(* Logix 5000 project; controller MV vendor 1 type 14 code 217 rev 31.11; software revision 31.00; part 52 of 53 *)
(* tags used below, declared in another part *)
   Alarm_Reset : BOOL;
   CWD : CHECKWORD_FLAGS;
   Default_Check_Time : DINT;
   Dummy : BOOL;
   Item_Faults_Are_Latched : BOOL;
   Item_Simulation_Flag : BOOL;
   Mike_050419 : BOOL;
   MV_data_file_address : INT;
   MV_data_file_value_to_move : DINT;
   MV_MV20R : PlantItem;   // MV20R
   MV_MV20R_ALARM : ALARM_DIGITAL;
   MV_MV20R_D : ALIAS FOR Remote_IO:14:O.Data.9;   // Rouser drive MV20
   MV_MV20R_R : ALIAS FOR Remote_IO:15:I.Data.25;   // MV20 Rouser running signal
   MV_MV21R : PlantItem;   // MV21R
   MV_MV21R_ALARM : ALARM_DIGITAL;
   MV_MV21R_D : ALIAS FOR Remote_IO:14:O.Data.10;   // Rouser drive MV21
   MV_MV21R_R : ALIAS FOR Remote_IO:15:I.Data.26;   // MV21 Rouser running signal
   MV_MV22R : PlantItem;   // MV22R
   MV_MV22R_ALARM : ALARM_DIGITAL;
   MV_MV22R_D : ALIAS FOR Remote_IO:14:O.Data.11;   // Rouser drive MV22
   MV_MV22R_R : ALIAS FOR Remote_IO:15:I.Data.27;   // MV22 Rouser running signal
   MV_MV23R : PlantItem;   // MV23R
   MV_MV23R_ALARM : ALARM_DIGITAL;
   MV_MV23R_D : ALIAS FOR Remote_IO:14:O.Data.12;   // Rouser drive MV23
   MV_MV23R_R : ALIAS FOR Remote_IO:15:I.Data.28;   // MV23 Rouser running signal
   MV_MV35R : PlantItem;   // MV35R
   MV_MV35R_ALARM : ALARM_DIGITAL;
   MV_MV35R_D : ALIAS FOR Remote_IO:14:O.Data.8;   // Rouser drive MV35
   MV_MV35R_R : ALIAS FOR Remote_IO:15:I.Data.24;   // MV35 Rouser running signal
   MV_N101 : INT[255];   // AT INT Fermentation control integer workspace
   MV_N105 : INT[255];   // ROUSE_CTRL Rouser control progr am working regs
   MV_N105_0_1_Output_Bit : BOOL;
   MV_N105_0_6_Output_Bit : BOOL;
   MV_N105_0_7_Output_Bit : BOOL;
   MV_N105_0_8_Output_Bit : BOOL;
   MV_N106 : INT[255];   // ROUSE_BUFF Rouser control vesse l data buffer
   MV_N110 : INT[255];   // MV DATA 0 CURRENT FV DATA
   MV_N111 : INT[50];   // MV 1, CURRENT FV DATA
   MV_N112 : INT[50];   // MV 2, CURRENT FV DATA
   MV_N113 : INT[50];   // MV 3, CURRENT FV DATA
   MV_N114 : INT[50];   // MV 4, CURRENT FV DATA
   MV_N115 : INT[50];   // MV 5, CURRENT FV DATA
   MV_N116 : INT[50];   // MV 6, CURRENT FV DATA
   MV_N117 : INT[50];   // MV 7, CURRENT FV DATA
   MV_N118 : INT[50];   // MV 8, CURRENT FV DATA
   MV_N119 : INT[50];   // MV 9, CURRENT FV DATA
   MV_N12 : INT[255];   // SYS_PARMS System Parameter Fil e
   MV_N120 : INT[50];   // MV 10, CURRENT FV DATA
   MV_N121 : INT[50];   // MV 11, CURRENT FV DATA
   MV_N122 : INT[50];   // MV 12, CURRENT FV DATA
   MV_N123 : INT[50];   // MV 13, CURRENT FV DATA
   MV_N124 : INT[50];   // MV 14, CURRENT FV DATA
   MV_N125 : INT[50];   // MV 15, CURRENT FV DATA
   MV_N126 : INT[50];   // MV 16, CURRENT FV DATA
   MV_N127 : INT[50];   // MV 17, CURRENT FV DATA
   MV_N128 : INT[50];   // MV 18, CURRENT FV DATA
   MV_N129 : INT[50];   // MV 19, CURRENT FV DATA
   MV_N130 : INT[50];   // MV 30, CURRENT FV DATA
   MV_N131 : INT[50];   // MV 31, CURRENT FV DATA
   MV_N132 : INT[50];   // MV 32, CURRENT FV DATA
   MV_N133 : INT[50];   // MV 33, CURRENT FV DATA
   MV_N134 : INT[50];   // MV 34, CURRENT FV DATA
   MV_N135 : INT[50];   // MV 35, CURRENT FV DATA
   MV_N136 : INT[50];   // MV 20, CURRENT FV DATA
   MV_N137 : INT[50];   // MV 21, CURRENT FV DATA
   MV_N138 : INT[50];   // MV 22, CURRENT FV DATA
   MV_N139 : INT[50];   // MV 23, CURRENT FV DATA
   MV_N140 : INT[50];   // MV 36, CURRENT FV DATA
   MV_N141 : INT[50];   // MV 37, CURRENT FV DATA
   MV_N142 : INT[50];   // MV 38, CURRENT FV DATA
   MV_N143 : INT[50];   // MV 39, CURRENT FV DATA
   MV_N144 : INT[50];   // MV 40, CURRENT FV DATA
   MV_N145 : INT[50];   // MV 41, CURRENT FV DATA
   MV_N146 : INT[50];   // MV 42, CURRENT FV DATA
   MV_N147 : INT[50];   // MV 43, CURRENT FV DATA
   MV_N148 : INT[50];   // MV 44, CURRENT FV DATA
   MV_N149 : INT[50];   // MV 45, CURRENT FV DATA
   MV_N150 : INT[50];   // MV 36, CURRENT FV DATA
   MV_N151 : INT[50];   // MV 47, CURRENT FV DATA
   MV_SFile : INT[255];   // SLC Equivalent System File, So Original Code Can Remain
   MV_T4 : TIMER[20];
   MV_value_to_set : INT;
   MV_word_offset : INT;
   One_Second_One_Scan : ALIAS FOR One_Second_1_scan;
   Scada_Pump_Fault_No : DINT;
   Scada_Pump_H_Fault_No : DINT;
   Scada_Pump_T_Fault_No : DINT;
   Unused_Healthy_Feedback : BOOL;
   Unused_NotTripped_Feedback : BOOL;
(* MV_Common, continued *)

   24: [NEQ(MV_MV35R.DriveBits,0) OTE(MV_MV35R.CW.[CWD.AUTODRV]) ,[XIC(MV_MV35R.CW.[CWD.AUTODRV]) XIO(MV_MV35R.CW.[CWD.MANUAL]) ,XIC(MV_MV35R.CW.[CWD.MANDRV]) XIC(MV_MV35R.CW.[CWD.MANUAL]) ] OTE(MV_MV35R.CW.[CWD.OUTPUT]) ,XIC(MV_MV35R.CW.[CWD.OUTPUT]) OTE(MV_MV35R_D) ,XIC(S:FS) [OTU(MV_MV35R.CW.[CWD.MANUAL]) ,LEQ(MV_MV35R.CheckTime,0) MOV(Default_Check_Time,MV_MV35R.CheckTime) ] ,[[XIC(MV_MV35R_R) XIO(Item_Simulation_Flag) ,XIC(Item_Simulation_Flag) [XIC(MV_MV35R.CW.[CWD.OUTPUT]) XIO(MV_MV35R.CW.[CWD.SIMFAIL]) ,XIO(MV_MV35R.CW.[CWD.OUTPUT]) XIC(MV_MV35R.CW.[CWD.SIMFAIL]) ] ] OTE(MV_MV35R.CW.[CWD.RUNFB]) ,[XIC(Item_Simulation_Flag) ,XIC(MV_MV35R.CW.[CWD.CHECKOFF]) ,XIC(Unused_Healthy_Feedback) ] OTE(MV_MV35R.CW.[CWD.HEALTHYFB]) ,[XIC(Item_Simulation_Flag) ,XIC(MV_MV35R.CW.[CWD.CHECKOFF]) ,XIC(Unused_NotTripped_Feedback) ] OTE(MV_MV35R.CW.[CWD.NOTTRIPPEDFB]) ] ,[XIC(MV_MV35R.CW.[CWD.AUTODRV]) XIO(MV_MV35R.CW.[CWD.PREVSCAN]) ,XIO(MV_MV35R.CW.[CWD.AUTODRV]) XIC(MV_MV35R.CW.[CWD.PREVSCAN]) ] CLR(MV_MV35R.CheckTimer) ,XIC(One_Second_One_Scan) LES(MV_MV35R.CheckTimer,MV_MV35R.CheckTime) ADD(MV_MV35R.CheckTimer,1,MV_MV35R.CheckTimer) ,XIO(MV_MV35R.CW.[CWD.FAULT]) OTU(MV_MV35R.CW.[CWD.FAULTLOGGED]) ,[GEQ(MV_MV35R.CheckTimer,MV_MV35R.CheckTime) [XIC(MV_MV35R.CW.[CWD.OUTPUT]) XIO(MV_MV35R.CW.[CWD.RUNFB]) ,XIO(MV_MV35R.CW.[CWD.OUTPUT]) XIC(MV_MV35R.CW.[CWD.RUNFB]) ] ,XIO(MV_MV35R.CW.[CWD.HEALTHYFB]) ,XIO(MV_MV35R.CW.[CWD.NOTTRIPPEDFB]) ,XIC(MV_MV35R.CW.[CWD.FAULT]) XIC(Item_Faults_Are_Latched) ,XIC(MV_MV35R.CW.[CWD.HIGHLIGHT]) ] XIO(MV_MV35R.CW.[CWD.CHECKOFF]) XIO(Alarm_Reset) [OTE(MV_MV35R.CW.[CWD.FAULT]) ,ALMD(MV_MV35R_ALARM,0,0,0,0) ] ,XIC(MV_MV35R.CW.[CWD.OUTPUT]) OTE(MV_MV35R.CW.[CWD.PREVSCAN]) ,XIC(MV_MV35R.CW.[CWD.FAULT]) EQU(Scada_Pump_Fault_No,0) XIO(MV_MV35R.CW.[CWD.FAULTLOGGED]) [MOV(20001,Scada_Pump_Fault_No) ,OTL(MV_MV35R.CW.[CWD.FAULTLOGGED]) ] ,XIO(MV_MV35R.CW.[CWD.HEALTHYFB]) EQU(Scada_Pump_H_Fault_No,0) XIO(MV_MV35R.CW.[CWD.HEALTHYFAULTLOGGED]) [MOV(20001,Scada_Pump_H_Fault_No) ,OTL(MV_MV35R.CW.[CWD.HEALTHYFAULTLOGGED]) ] ,XIO(MV_MV35R.CW.[CWD.NOTTRIPPEDFB]) EQU(Scada_Pump_H_Fault_No,0) XIO(MV_MV35R.CW.[CWD.TRIPPEDFAULTLOGGED]) [MOV(20001,Scada_Pump_T_Fault_No) ,OTL(MV_MV35R.CW.[CWD.TRIPPEDFAULTLOGGED]) ] ];
   25: [NEQ(MV_MV20R.DriveBits,0) OTE(MV_MV20R.CW.[CWD.AUTODRV]) ,[XIC(MV_MV20R.CW.[CWD.AUTODRV]) XIO(MV_MV20R.CW.[CWD.MANUAL]) ,XIC(MV_MV20R.CW.[CWD.MANDRV]) XIC(MV_MV20R.CW.[CWD.MANUAL]) ] OTE(MV_MV20R.CW.[CWD.OUTPUT]) ,XIC(MV_MV20R.CW.[CWD.OUTPUT]) OTE(MV_MV20R_D) ,XIC(S:FS) [OTU(MV_MV20R.CW.[CWD.MANUAL]) ,LEQ(MV_MV20R.CheckTime,0) MOV(Default_Check_Time,MV_MV20R.CheckTime) ] ,[[XIC(MV_MV20R_R) XIO(Item_Simulation_Flag) ,XIC(Item_Simulation_Flag) [XIC(MV_MV20R.CW.[CWD.OUTPUT]) XIO(MV_MV20R.CW.[CWD.SIMFAIL]) ,XIO(MV_MV20R.CW.[CWD.OUTPUT]) XIC(MV_MV20R.CW.[CWD.SIMFAIL]) ] ] OTE(MV_MV20R.CW.[CWD.RUNFB]) ,[XIC(Item_Simulation_Flag) ,XIC(MV_MV20R.CW.[CWD.CHECKOFF]) ,XIC(Unused_Healthy_Feedback) ] OTE(MV_MV20R.CW.[CWD.HEALTHYFB]) ,[XIC(Item_Simulation_Flag) ,XIC(MV_MV20R.CW.[CWD.CHECKOFF]) ,XIC(Unused_NotTripped_Feedback) ] OTE(MV_MV20R.CW.[CWD.NOTTRIPPEDFB]) ] ,[XIC(MV_MV20R.CW.[CWD.AUTODRV]) XIO(MV_MV20R.CW.[CWD.PREVSCAN]) ,XIO(MV_MV20R.CW.[CWD.AUTODRV]) XIC(MV_MV20R.CW.[CWD.PREVSCAN]) ] CLR(MV_MV20R.CheckTimer) ,XIC(One_Second_One_Scan) LES(MV_MV20R.CheckTimer,MV_MV20R.CheckTime) ADD(MV_MV20R.CheckTimer,1,MV_MV20R.CheckTimer) ,XIO(MV_MV20R.CW.[CWD.FAULT]) OTU(MV_MV20R.CW.[CWD.FAULTLOGGED]) ,[GEQ(MV_MV20R.CheckTimer,MV_MV20R.CheckTime) [XIC(MV_MV20R.CW.[CWD.OUTPUT]) XIO(MV_MV20R.CW.[CWD.RUNFB]) ,XIO(MV_MV20R.CW.[CWD.OUTPUT]) XIC(MV_MV20R.CW.[CWD.RUNFB]) ] ,XIO(MV_MV20R.CW.[CWD.HEALTHYFB]) ,XIO(MV_MV20R.CW.[CWD.NOTTRIPPEDFB]) ,XIC(MV_MV20R.CW.[CWD.FAULT]) XIC(Item_Faults_Are_Latched) ,XIC(MV_MV20R.CW.[CWD.HIGHLIGHT]) ] XIO(MV_MV20R.CW.[CWD.CHECKOFF]) XIO(Alarm_Reset) [OTE(MV_MV20R.CW.[CWD.FAULT]) ,ALMD(MV_MV20R_ALARM,0,0,0,0) ] ,XIC(MV_MV20R.CW.[CWD.OUTPUT]) OTE(MV_MV20R.CW.[CWD.PREVSCAN]) ,XIC(MV_MV20R.CW.[CWD.FAULT]) EQU(Scada_Pump_Fault_No,0) XIO(MV_MV20R.CW.[CWD.FAULTLOGGED]) [MOV(20001,Scada_Pump_Fault_No) ,OTL(MV_MV20R.CW.[CWD.FAULTLOGGED]) ] ,XIO(MV_MV20R.CW.[CWD.HEALTHYFB]) EQU(Scada_Pump_H_Fault_No,0) XIO(MV_MV20R.CW.[CWD.HEALTHYFAULTLOGGED]) [MOV(20001,Scada_Pump_H_Fault_No) ,OTL(MV_MV20R.CW.[CWD.HEALTHYFAULTLOGGED]) ] ,XIO(MV_MV20R.CW.[CWD.NOTTRIPPEDFB]) EQU(Scada_Pump_H_Fault_No,0) XIO(MV_MV20R.CW.[CWD.TRIPPEDFAULTLOGGED]) [MOV(20001,Scada_Pump_T_Fault_No) ,OTL(MV_MV20R.CW.[CWD.TRIPPEDFAULTLOGGED]) ] ];
   26: [NEQ(MV_MV21R.DriveBits,0) OTE(MV_MV21R.CW.[CWD.AUTODRV]) ,[XIC(MV_MV21R.CW.[CWD.AUTODRV]) XIO(MV_MV21R.CW.[CWD.MANUAL]) ,XIC(MV_MV21R.CW.[CWD.MANDRV]) XIC(MV_MV21R.CW.[CWD.MANUAL]) ] OTE(MV_MV21R.CW.[CWD.OUTPUT]) ,XIC(MV_MV21R.CW.[CWD.OUTPUT]) OTE(MV_MV21R_D) ,XIC(S:FS) [OTU(MV_MV21R.CW.[CWD.MANUAL]) ,LEQ(MV_MV21R.CheckTime,0) MOV(Default_Check_Time,MV_MV21R.CheckTime) ] ,[[XIC(MV_MV21R_R) XIO(Item_Simulation_Flag) ,XIC(Item_Simulation_Flag) [XIC(MV_MV21R.CW.[CWD.OUTPUT]) XIO(MV_MV21R.CW.[CWD.SIMFAIL]) ,XIO(MV_MV21R.CW.[CWD.OUTPUT]) XIC(MV_MV21R.CW.[CWD.SIMFAIL]) ] ] OTE(MV_MV21R.CW.[CWD.RUNFB]) ,[XIC(Item_Simulation_Flag) ,XIC(MV_MV21R.CW.[CWD.CHECKOFF]) ,XIC(Unused_Healthy_Feedback) ] OTE(MV_MV21R.CW.[CWD.HEALTHYFB]) ,[XIC(Item_Simulation_Flag) ,XIC(MV_MV21R.CW.[CWD.CHECKOFF]) ,XIC(Unused_NotTripped_Feedback) ] OTE(MV_MV21R.CW.[CWD.NOTTRIPPEDFB]) ] ,[XIC(MV_MV21R.CW.[CWD.AUTODRV]) XIO(MV_MV21R.CW.[CWD.PREVSCAN]) ,XIO(MV_MV21R.CW.[CWD.AUTODRV]) XIC(MV_MV21R.CW.[CWD.PREVSCAN]) ] CLR(MV_MV21R.CheckTimer) ,XIC(One_Second_One_Scan) LES(MV_MV21R.CheckTimer,MV_MV21R.CheckTime) ADD(MV_MV21R.CheckTimer,1,MV_MV21R.CheckTimer) ,XIO(MV_MV21R.CW.[CWD.FAULT]) OTU(MV_MV21R.CW.[CWD.FAULTLOGGED]) ,[GEQ(MV_MV21R.CheckTimer,MV_MV21R.CheckTime) [XIC(MV_MV21R.CW.[CWD.OUTPUT]) XIO(MV_MV21R.CW.[CWD.RUNFB]) ,XIO(MV_MV21R.CW.[CWD.OUTPUT]) XIC(MV_MV21R.CW.[CWD.RUNFB]) ] ,XIO(MV_MV21R.CW.[CWD.HEALTHYFB]) ,XIO(MV_MV21R.CW.[CWD.NOTTRIPPEDFB]) ,XIC(MV_MV21R.CW.[CWD.FAULT]) XIC(Item_Faults_Are_Latched) ,XIC(MV_MV21R.CW.[CWD.HIGHLIGHT]) ] XIO(MV_MV21R.CW.[CWD.CHECKOFF]) XIO(Alarm_Reset) [OTE(MV_MV21R.CW.[CWD.FAULT]) ,ALMD(MV_MV21R_ALARM,0,0,0,0) ] ,XIC(MV_MV21R.CW.[CWD.OUTPUT]) OTE(MV_MV21R.CW.[CWD.PREVSCAN]) ,XIC(MV_MV21R.CW.[CWD.FAULT]) EQU(Scada_Pump_Fault_No,0) XIO(MV_MV21R.CW.[CWD.FAULTLOGGED]) [MOV(20001,Scada_Pump_Fault_No) ,OTL(MV_MV21R.CW.[CWD.FAULTLOGGED]) ] ,XIO(MV_MV21R.CW.[CWD.HEALTHYFB]) EQU(Scada_Pump_H_Fault_No,0) XIO(MV_MV21R.CW.[CWD.HEALTHYFAULTLOGGED]) [MOV(20001,Scada_Pump_H_Fault_No) ,OTL(MV_MV21R.CW.[CWD.HEALTHYFAULTLOGGED]) ] ,XIO(MV_MV21R.CW.[CWD.NOTTRIPPEDFB]) EQU(Scada_Pump_H_Fault_No,0) XIO(MV_MV21R.CW.[CWD.TRIPPEDFAULTLOGGED]) [MOV(20001,Scada_Pump_T_Fault_No) ,OTL(MV_MV21R.CW.[CWD.TRIPPEDFAULTLOGGED]) ] ];
   27: [NEQ(MV_MV22R.DriveBits,0) OTE(MV_MV22R.CW.[CWD.AUTODRV]) ,[XIC(MV_MV22R.CW.[CWD.AUTODRV]) XIO(MV_MV22R.CW.[CWD.MANUAL]) ,XIC(MV_MV22R.CW.[CWD.MANDRV]) XIC(MV_MV22R.CW.[CWD.MANUAL]) ] OTE(MV_MV22R.CW.[CWD.OUTPUT]) ,XIC(MV_MV22R.CW.[CWD.OUTPUT]) OTE(MV_MV22R_D) ,XIC(S:FS) [OTU(MV_MV22R.CW.[CWD.MANUAL]) ,LEQ(MV_MV22R.CheckTime,0) MOV(Default_Check_Time,MV_MV22R.CheckTime) ] ,[[XIC(MV_MV22R_R) XIO(Item_Simulation_Flag) ,XIC(Item_Simulation_Flag) [XIC(MV_MV22R.CW.[CWD.OUTPUT]) XIO(MV_MV22R.CW.[CWD.SIMFAIL]) ,XIO(MV_MV22R.CW.[CWD.OUTPUT]) XIC(MV_MV22R.CW.[CWD.SIMFAIL]) ] ] OTE(MV_MV22R.CW.[CWD.RUNFB]) ,[XIC(Item_Simulation_Flag) ,XIC(MV_MV22R.CW.[CWD.CHECKOFF]) ,XIC(Unused_Healthy_Feedback) ] OTE(MV_MV22R.CW.[CWD.HEALTHYFB]) ,[XIC(Item_Simulation_Flag) ,XIC(MV_MV22R.CW.[CWD.CHECKOFF]) ,XIC(Unused_NotTripped_Feedback) ] OTE(MV_MV22R.CW.[CWD.NOTTRIPPEDFB]) ] ,[XIC(MV_MV22R.CW.[CWD.AUTODRV]) XIO(MV_MV22R.CW.[CWD.PREVSCAN]) ,XIO(MV_MV22R.CW.[CWD.AUTODRV]) XIC(MV_MV22R.CW.[CWD.PREVSCAN]) ] CLR(MV_MV22R.CheckTimer) ,XIC(One_Second_One_Scan) LES(MV_MV22R.CheckTimer,MV_MV22R.CheckTime) ADD(MV_MV22R.CheckTimer,1,MV_MV22R.CheckTimer) ,XIO(MV_MV22R.CW.[CWD.FAULT]) OTU(MV_MV22R.CW.[CWD.FAULTLOGGED]) ,[GEQ(MV_MV22R.CheckTimer,MV_MV22R.CheckTime) [XIC(MV_MV22R.CW.[CWD.OUTPUT]) XIO(MV_MV22R.CW.[CWD.RUNFB]) ,XIO(MV_MV22R.CW.[CWD.OUTPUT]) XIC(MV_MV22R.CW.[CWD.RUNFB]) ] ,XIO(MV_MV22R.CW.[CWD.HEALTHYFB]) ,XIO(MV_MV22R.CW.[CWD.NOTTRIPPEDFB]) ,XIC(MV_MV22R.CW.[CWD.FAULT]) XIC(Item_Faults_Are_Latched) ,XIC(MV_MV22R.CW.[CWD.HIGHLIGHT]) ] XIO(MV_MV22R.CW.[CWD.CHECKOFF]) XIO(Alarm_Reset) [OTE(MV_MV22R.CW.[CWD.FAULT]) ,ALMD(MV_MV22R_ALARM,0,0,0,0) ] ,XIC(MV_MV22R.CW.[CWD.OUTPUT]) OTE(MV_MV22R.CW.[CWD.PREVSCAN]) ,XIC(MV_MV22R.CW.[CWD.FAULT]) EQU(Scada_Pump_Fault_No,0) XIO(MV_MV22R.CW.[CWD.FAULTLOGGED]) [MOV(20001,Scada_Pump_Fault_No) ,OTL(MV_MV22R.CW.[CWD.FAULTLOGGED]) ] ,XIO(MV_MV22R.CW.[CWD.HEALTHYFB]) EQU(Scada_Pump_H_Fault_No,0) XIO(MV_MV22R.CW.[CWD.HEALTHYFAULTLOGGED]) [MOV(20001,Scada_Pump_H_Fault_No) ,OTL(MV_MV22R.CW.[CWD.HEALTHYFAULTLOGGED]) ] ,XIO(MV_MV22R.CW.[CWD.NOTTRIPPEDFB]) EQU(Scada_Pump_H_Fault_No,0) XIO(MV_MV22R.CW.[CWD.TRIPPEDFAULTLOGGED]) [MOV(20001,Scada_Pump_T_Fault_No) ,OTL(MV_MV22R.CW.[CWD.TRIPPEDFAULTLOGGED]) ] ];
   28: [NEQ(MV_MV23R.DriveBits,0) OTE(MV_MV23R.CW.[CWD.AUTODRV]) ,[XIC(MV_MV23R.CW.[CWD.AUTODRV]) XIO(MV_MV23R.CW.[CWD.MANUAL]) ,XIC(MV_MV23R.CW.[CWD.MANDRV]) XIC(MV_MV23R.CW.[CWD.MANUAL]) ] OTE(MV_MV23R.CW.[CWD.OUTPUT]) ,XIC(MV_MV23R.CW.[CWD.OUTPUT]) OTE(MV_MV23R_D) ,XIC(S:FS) [OTU(MV_MV23R.CW.[CWD.MANUAL]) ,LEQ(MV_MV23R.CheckTime,0) MOV(Default_Check_Time,MV_MV23R.CheckTime) ] ,[[XIC(MV_MV23R_R) XIO(Item_Simulation_Flag) ,XIC(Item_Simulation_Flag) [XIC(MV_MV23R.CW.[CWD.OUTPUT]) XIO(MV_MV23R.CW.[CWD.SIMFAIL]) ,XIO(MV_MV23R.CW.[CWD.OUTPUT]) XIC(MV_MV23R.CW.[CWD.SIMFAIL]) ] ] OTE(MV_MV23R.CW.[CWD.RUNFB]) ,[XIC(Item_Simulation_Flag) ,XIC(MV_MV23R.CW.[CWD.CHECKOFF]) ,XIC(Unused_Healthy_Feedback) ] OTE(MV_MV23R.CW.[CWD.HEALTHYFB]) ,[XIC(Item_Simulation_Flag) ,XIC(MV_MV23R.CW.[CWD.CHECKOFF]) ,XIC(Unused_NotTripped_Feedback) ] OTE(MV_MV23R.CW.[CWD.NOTTRIPPEDFB]) ] ,[XIC(MV_MV23R.CW.[CWD.AUTODRV]) XIO(MV_MV23R.CW.[CWD.PREVSCAN]) ,XIO(MV_MV23R.CW.[CWD.AUTODRV]) XIC(MV_MV23R.CW.[CWD.PREVSCAN]) ] CLR(MV_MV23R.CheckTimer) ,XIC(One_Second_One_Scan) LES(MV_MV23R.CheckTimer,MV_MV23R.CheckTime) ADD(MV_MV23R.CheckTimer,1,MV_MV23R.CheckTimer) ,XIO(MV_MV23R.CW.[CWD.FAULT]) OTU(MV_MV23R.CW.[CWD.FAULTLOGGED]) ,[GEQ(MV_MV23R.CheckTimer,MV_MV23R.CheckTime) [XIC(MV_MV23R.CW.[CWD.OUTPUT]) XIO(MV_MV23R.CW.[CWD.RUNFB]) ,XIO(MV_MV23R.CW.[CWD.OUTPUT]) XIC(MV_MV23R.CW.[CWD.RUNFB]) ] ,XIO(MV_MV23R.CW.[CWD.HEALTHYFB]) ,XIO(MV_MV23R.CW.[CWD.NOTTRIPPEDFB]) ,XIC(MV_MV23R.CW.[CWD.FAULT]) XIC(Item_Faults_Are_Latched) ,XIC(MV_MV23R.CW.[CWD.HIGHLIGHT]) ] XIO(MV_MV23R.CW.[CWD.CHECKOFF]) XIO(Alarm_Reset) [OTE(MV_MV23R.CW.[CWD.FAULT]) ,ALMD(MV_MV23R_ALARM,0,0,0,0) ] ,XIC(MV_MV23R.CW.[CWD.OUTPUT]) OTE(MV_MV23R.CW.[CWD.PREVSCAN]) ,XIC(MV_MV23R.CW.[CWD.FAULT]) EQU(Scada_Pump_Fault_No,0) XIO(MV_MV23R.CW.[CWD.FAULTLOGGED]) [MOV(20001,Scada_Pump_Fault_No) ,OTL(MV_MV23R.CW.[CWD.FAULTLOGGED]) ] ,XIO(MV_MV23R.CW.[CWD.HEALTHYFB]) EQU(Scada_Pump_H_Fault_No,0) XIO(MV_MV23R.CW.[CWD.HEALTHYFAULTLOGGED]) [MOV(20001,Scada_Pump_H_Fault_No) ,OTL(MV_MV23R.CW.[CWD.HEALTHYFAULTLOGGED]) ] ,XIO(MV_MV23R.CW.[CWD.NOTTRIPPEDFB]) EQU(Scada_Pump_H_Fault_No,0) XIO(MV_MV23R.CW.[CWD.TRIPPEDFAULTLOGGED]) [MOV(20001,Scada_Pump_T_Fault_No) ,OTL(MV_MV23R.CW.[CWD.TRIPPEDFAULTLOGGED]) ] ];
END_ROUTINE

ROUTINE MV_ROUSERS_110   (* ladder *)
   // If PC has requested timed rouser operation save current rouser mode and load rousing time
   0: [LIM(29,MV_N105[2],56) ,EQU(MV_N105[2],94) ,LIM(336,MV_N105[2],347) ][ADD(MV_N105[2],82,MV_N105[4]) ,EQU(MV_N105[2],94) MOV(139,MV_N105[4]) ,LIM(336,MV_N105[2],347) SUB(MV_N105[2],196,MV_N105[4]) ,JSR(MV_Set_FV_Datafile_Value,3,MV_N105[3],MV_N105[4],31) ,JSR(MV_Get_FV_Datafile_Value,2,MV_N105[4],32) JSR(MV_Set_FV_Datafile_Value,3,MV_data_file_value_to_move,MV_N105[4],34) ,JSR(MV_Set_FV_Datafile_Value,3,3,MV_N105[4],32) ,CLR(MV_N105[2]) ];
   // Set pointer to first vessel data file at power up
   1: XIC(S:FS)OSR(MV_N105[0].1,MV_N105_0_1_Output_Bit)XIC(MV_N105_0_1_Output_Bit)MOV(111,MV_N105[1]);
   // Trigger rouser daily operation if current time equals time in settings file N12
   2: EQU(MV_SFile[40],MV_N12[1])EQU(MV_SFile[41],MV_N12[2])EQU(MV_SFile[42],0)OSR(MV_N105[0].6,MV_N105_0_6_Output_Bit)XIC(MV_N105_0_6_Output_Bit)OTL(MV_N105[0].2);
   // Set daily rousing latch when vessel loop at 1st vessel
   3: XIC(MV_N105[0].2)EQU(MV_N105[1],111)[OTL(MV_N105[0].3) ,OTU(MV_N105[0].2) ];
   // Trigger rouser hourly operation if current time equals time in settings file N12
   4: EQU(MV_SFile[41],0)EQU(MV_SFile[42],0)OSR(MV_N105[0].8,MV_N105_0_8_Output_Bit)XIC(MV_N105_0_8_Output_Bit)OTL(MV_N105[0].9);
   // Set hourly rousing latch when vessel loop at 1st vessel
   5: XIC(MV_N105[0].9)EQU(MV_N105[1],111)[OTL(MV_N105[0].10) ,OTU(MV_N105[0].9) ];
   // Inform rouser loop one minute has elapsed
   6: EQU(MV_SFile[42],0)OSR(MV_N105[0].7,MV_N105_0_7_Output_Bit)XIC(MV_N105_0_7_Output_Bit)OTL(MV_N105[0].4);
   7: XIC(MV_N105[0].4)EQU(MV_N105[1],111)[OTL(MV_N105[0].0) ,OTU(MV_N105[0].4) ];
   // ROUSER CONTROL LOOP RUN CONTINUOUSLY BUT SEPARATES VESSELS BY 1 SEC
   8: XIC(MV_N105[0].0)XIC(MV_T4[2].DN)MCR();
   // Take copy of current vessel data file
   9: JSR(MV_Copy_Vessel_File,2,MV_N105[1],106);
   // If elapsed time > 2 hours enable rouser
   10: LIM(8,MV_N106[24],16)[GEQ(MV_N106[27],20) OTL(MV_N106[15].7) ,LES(MV_N106[27],20) OTU(MV_N106[15].7) ];
   11: XIC(Mike_050419)NEQ(MV_N106[32],3)EQU(MV_N105[1],MV_N105[1])MOV(MV_N106[32],MV_N106[34]);
   // If time remains for timed rouser operation and one minute has elapsed decrement by 1 minute
   12: GRT(MV_N106[31],0)XIC(MV_N105[0].0)[SUB(MV_N106[31],1,MV_N106[31]) ,XIC(Mike_050419) LEQ(MV_N106[31],0) MOV(MV_N106[34],MV_N106[32]) ];
   // Restore rouser mode of operation after timed rouse operation completes
   13: XIO(Mike_050419)EQU(MV_N106[32],3)LEQ(MV_N106[31],0)MOV(MV_N106[34],MV_N106[32]);
   // If it is time to do daily rouse load daily rousing duration to timed operation timer
   14: XIC(MV_N105[0].3)EQU(MV_N106[32],2)XIO(MV_N106[29].1)MOV(MV_N12[3],MV_N106[31]);
   // If it is time to do hourly rouse load hourly rousing duration to timed operation timer
   15: XIC(MV_N105[0].10)EQU(MV_N106[32],4)XIO(MV_N106[29].1)MOV(MV_N12[4],MV_N106[31]);
   // Calculate temperature at which rouser is to operate
   16: ADD(MV_N106[26],3,MV_N101[9]);
   // If actual temperature > setpoint + 0.3 degC set flag for rousing required
   17: GRT(MV_N106[25],MV_N101[9])NEQ(MV_N106[24],0)OTE(MV_N106[30].2);
   // Set flag to request rouser to run as required
   18: [XIC(MV_N106[15].7) ,LIM(140,MV_N105[1],151) ]NEQ(MV_N106[32],0)[GRT(MV_N106[31],0) ,EQU(MV_N106[32],1) ,[XIC(MV_N106[30].0) ,XIC(MV_N106[30].2) ] XIO(MV_N106[29].1) ]OTE(MV_N106[30].1);
   // Save vessel data file
   19: JSR(MV_Copy_Vessel_File,2,106,MV_N105[1]);
   // Next vessel
   20: ADD(MV_N105[1],1,MV_N105[1]);
   // If all vessels done restart loop operation from 1st vessel
   21: GRT(MV_N105[1],151)[MOV(111,MV_N105[1]) ,OTU(MV_N105[0].0) ,OTU(MV_N105[0].3) ,OTU(MV_N105[0].10) ];
   22: MCR();
END_ROUTINE

ROUTINE MV_Set_FV_Datafile_Value   (* ladder *)
   // Routine to Set the value of something within the FV Data Files, Used to replace indirection originally used
   0: SBR(MV_value_to_set,MV_data_file_address,MV_word_offset)OTE(Dummy);
   1: EQU(MV_data_file_address,106)MOV(MV_value_to_set,MV_N106[MV_word_offset]);
   2: EQU(MV_data_file_address,110)MOV(MV_value_to_set,MV_N110[MV_word_offset]);
   3: EQU(MV_data_file_address,111)MOV(MV_value_to_set,MV_N111[MV_word_offset]);
   4: EQU(MV_data_file_address,112)MOV(MV_value_to_set,MV_N112[MV_word_offset]);
   5: EQU(MV_data_file_address,113)MOV(MV_value_to_set,MV_N113[MV_word_offset]);
   6: EQU(MV_data_file_address,114)MOV(MV_value_to_set,MV_N114[MV_word_offset]);
   7: EQU(MV_data_file_address,115)MOV(MV_value_to_set,MV_N115[MV_word_offset]);
   8: EQU(MV_data_file_address,116)MOV(MV_value_to_set,MV_N116[MV_word_offset]);
   9: EQU(MV_data_file_address,117)MOV(MV_value_to_set,MV_N117[MV_word_offset]);
   10: EQU(MV_data_file_address,118)MOV(MV_value_to_set,MV_N118[MV_word_offset]);
   11: EQU(MV_data_file_address,119)MOV(MV_value_to_set,MV_N119[MV_word_offset]);
   12: EQU(MV_data_file_address,120)MOV(MV_value_to_set,MV_N120[MV_word_offset]);
   13: EQU(MV_data_file_address,121)MOV(MV_value_to_set,MV_N121[MV_word_offset]);
   14: EQU(MV_data_file_address,122)MOV(MV_value_to_set,MV_N122[MV_word_offset]);
   15: EQU(MV_data_file_address,123)MOV(MV_value_to_set,MV_N123[MV_word_offset]);
   16: EQU(MV_data_file_address,124)MOV(MV_value_to_set,MV_N124[MV_word_offset]);
   17: EQU(MV_data_file_address,125)MOV(MV_value_to_set,MV_N125[MV_word_offset]);
   18: EQU(MV_data_file_address,126)MOV(MV_value_to_set,MV_N126[MV_word_offset]);
   19: EQU(MV_data_file_address,127)MOV(MV_value_to_set,MV_N127[MV_word_offset]);
   20: EQU(MV_data_file_address,128)MOV(MV_value_to_set,MV_N128[MV_word_offset]);
   21: EQU(MV_data_file_address,129)MOV(MV_value_to_set,MV_N129[MV_word_offset]);
   22: EQU(MV_data_file_address,130)MOV(MV_value_to_set,MV_N130[MV_word_offset]);
   23: EQU(MV_data_file_address,131)MOV(MV_value_to_set,MV_N131[MV_word_offset]);
   24: EQU(MV_data_file_address,132)MOV(MV_value_to_set,MV_N132[MV_word_offset]);
   25: EQU(MV_data_file_address,133)MOV(MV_value_to_set,MV_N133[MV_word_offset]);
   26: EQU(MV_data_file_address,134)MOV(MV_value_to_set,MV_N134[MV_word_offset]);
   27: EQU(MV_data_file_address,135)MOV(MV_value_to_set,MV_N135[MV_word_offset]);
   28: EQU(MV_data_file_address,136)MOV(MV_value_to_set,MV_N136[MV_word_offset]);
   29: EQU(MV_data_file_address,137)MOV(MV_value_to_set,MV_N137[MV_word_offset]);
   30: EQU(MV_data_file_address,138)MOV(MV_value_to_set,MV_N138[MV_word_offset]);
   31: EQU(MV_data_file_address,139)MOV(MV_value_to_set,MV_N139[MV_word_offset]);
   32: EQU(MV_data_file_address,140)MOV(MV_value_to_set,MV_N140[MV_word_offset]);
   33: EQU(MV_data_file_address,141)MOV(MV_value_to_set,MV_N141[MV_word_offset]);
   34: EQU(MV_data_file_address,142)MOV(MV_value_to_set,MV_N142[MV_word_offset]);
   35: EQU(MV_data_file_address,143)MOV(MV_value_to_set,MV_N143[MV_word_offset]);
   36: EQU(MV_data_file_address,144)MOV(MV_value_to_set,MV_N144[MV_word_offset]);
   37: EQU(MV_data_file_address,145)MOV(MV_value_to_set,MV_N145[MV_word_offset]);
   38: EQU(MV_data_file_address,146)MOV(MV_value_to_set,MV_N146[MV_word_offset]);
   39: EQU(MV_data_file_address,147)MOV(MV_value_to_set,MV_N147[MV_word_offset]);
   40: EQU(MV_data_file_address,148)MOV(MV_value_to_set,MV_N148[MV_word_offset]);
   41: EQU(MV_data_file_address,149)MOV(MV_value_to_set,MV_N149[MV_word_offset]);
   42: EQU(MV_data_file_address,150)MOV(MV_value_to_set,MV_N150[MV_word_offset]);
   43: EQU(MV_data_file_address,151)MOV(MV_value_to_set,MV_N151[MV_word_offset]);
   44: RET();
END_ROUTINE
